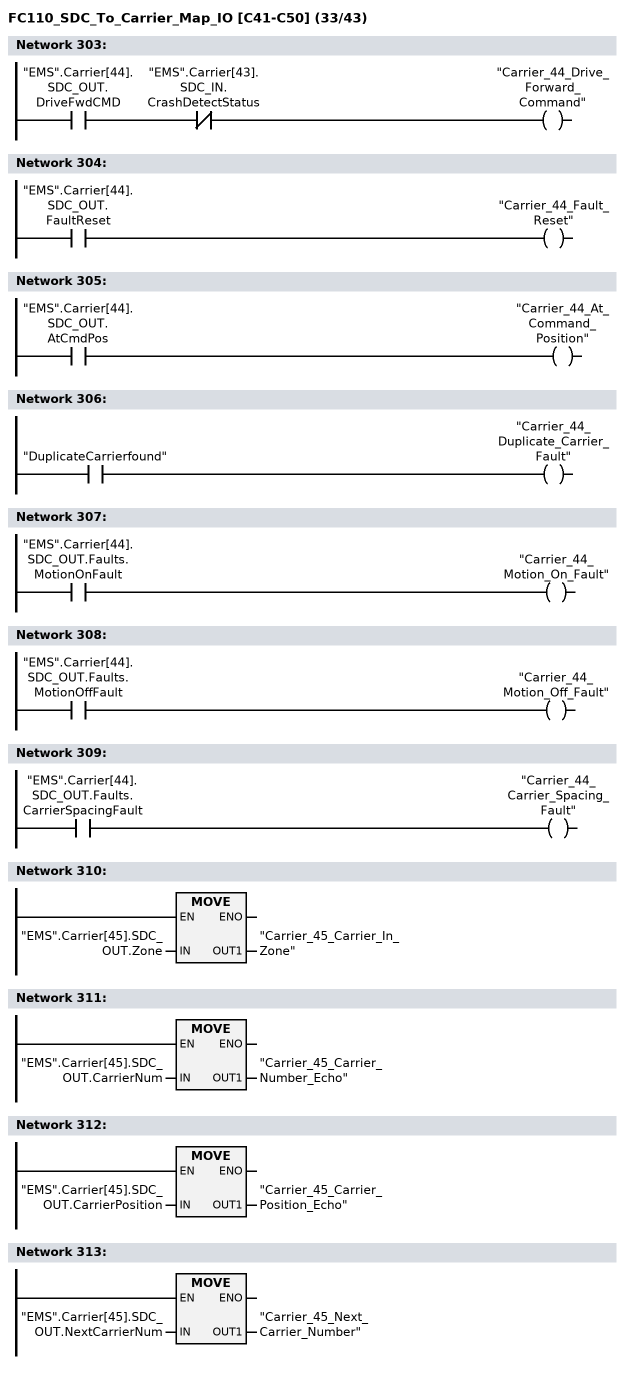
   RUNG wire#powerrail
      Contact( "EMS".Carrier[44].SDC_OUT.DriveFwdCMD )
      I_Contact( "EMS".Carrier[43].SDC_IN.CrashDetectStatus )
      Coil( "Carrier_44_Drive_Forward_Command" )
   END_RUNG
   // the same network as SCL:
   "Carrier_44_Drive_Forward_Command" := "EMS".Carrier[44].SDC_OUT.DriveFwdCMD AND NOT "EMS".Carrier[43].SDC_IN.CrashDetectStatus;
END_REGION

REGION Network 304
   RUNG wire#powerrail
      Contact( "EMS".Carrier[44].SDC_OUT.FaultReset )
      Coil( "Carrier_44_Fault_Reset" )
   END_RUNG
   // the same network as SCL:
   "Carrier_44_Fault_Reset" := "EMS".Carrier[44].SDC_OUT.FaultReset;
END_REGION

REGION Network 305
   RUNG wire#powerrail
      Contact( "EMS".Carrier[44].SDC_OUT.AtCmdPos )
      Coil( "Carrier_44_At_Command_Position" )
   END_RUNG
   // the same network as SCL:
   "Carrier_44_At_Command_Position" := "EMS".Carrier[44].SDC_OUT.AtCmdPos;
END_REGION

REGION Network 306
   RUNG wire#powerrail
      Contact( "DuplicateCarrierfound" )
      Coil( "Carrier_44_Duplicate_Carrier_Fault" )
   END_RUNG
   // the same network as SCL:
   "Carrier_44_Duplicate_Carrier_Fault" := "DuplicateCarrierfound";
END_REGION

REGION Network 307
   RUNG wire#powerrail
      Contact( "EMS".Carrier[44].SDC_OUT.Faults.MotionOnFault )
      Coil( "Carrier_44_Motion_On_Fault" )
   END_RUNG
   // the same network as SCL:
   "Carrier_44_Motion_On_Fault" := "EMS".Carrier[44].SDC_OUT.Faults.MotionOnFault;
END_REGION

REGION Network 308
   RUNG wire#powerrail
      Contact( "EMS".Carrier[44].SDC_OUT.Faults.MotionOffFault )
      Coil( "Carrier_44_Motion_Off_Fault" )
   END_RUNG
   // the same network as SCL:
   "Carrier_44_Motion_Off_Fault" := "EMS".Carrier[44].SDC_OUT.Faults.MotionOffFault;
END_REGION

REGION Network 309
   RUNG wire#powerrail
      Contact( "EMS".Carrier[44].SDC_OUT.Faults.CarrierSpacingFault )
      Coil( "Carrier_44_Carrier_Spacing_Fault" )
   END_RUNG
   // the same network as SCL:
   "Carrier_44_Carrier_Spacing_Fault" := "EMS".Carrier[44].SDC_OUT.Faults.CarrierSpacingFault;
END_REGION

REGION Network 310
   RUNG wire#powerrail
      Move(in := "EMS".Carrier[45].SDC_OUT.Zone, out1 => "Carrier_45_Carrier_In_Zone")
   END_RUNG
   // the same network as SCL:
   "Carrier_45_Carrier_In_Zone" := "EMS".Carrier[45].SDC_OUT.Zone;
END_REGION

REGION Network 311
   RUNG wire#powerrail
      Move(in := "EMS".Carrier[45].SDC_OUT.CarrierNum, out1 => "Carrier_45_Carrier_Number_Echo")
   END_RUNG
   // the same network as SCL:
   "Carrier_45_Carrier_Number_Echo" := "EMS".Carrier[45].SDC_OUT.CarrierNum;
END_REGION

REGION Network 312
   RUNG wire#powerrail
      Move(in := "EMS".Carrier[45].SDC_OUT.CarrierPosition, out1 => "Carrier_45_Carrier_Position_Echo")
   END_RUNG
   // the same network as SCL:
   "Carrier_45_Carrier_Position_Echo" := "EMS".Carrier[45].SDC_OUT.CarrierPosition;
END_REGION

REGION Network 313
   RUNG wire#powerrail
      Move(in := "EMS".Carrier[45].SDC_OUT.NextCarrierNum, out1 => "Carrier_45_Next_Carrier_Number")
   END_RUNG
   // the same network as SCL:
   "Carrier_45_Next_Carrier_Number" := "EMS".Carrier[45].SDC_OUT.NextCarrierNum;
END_REGION

REGION Network 314
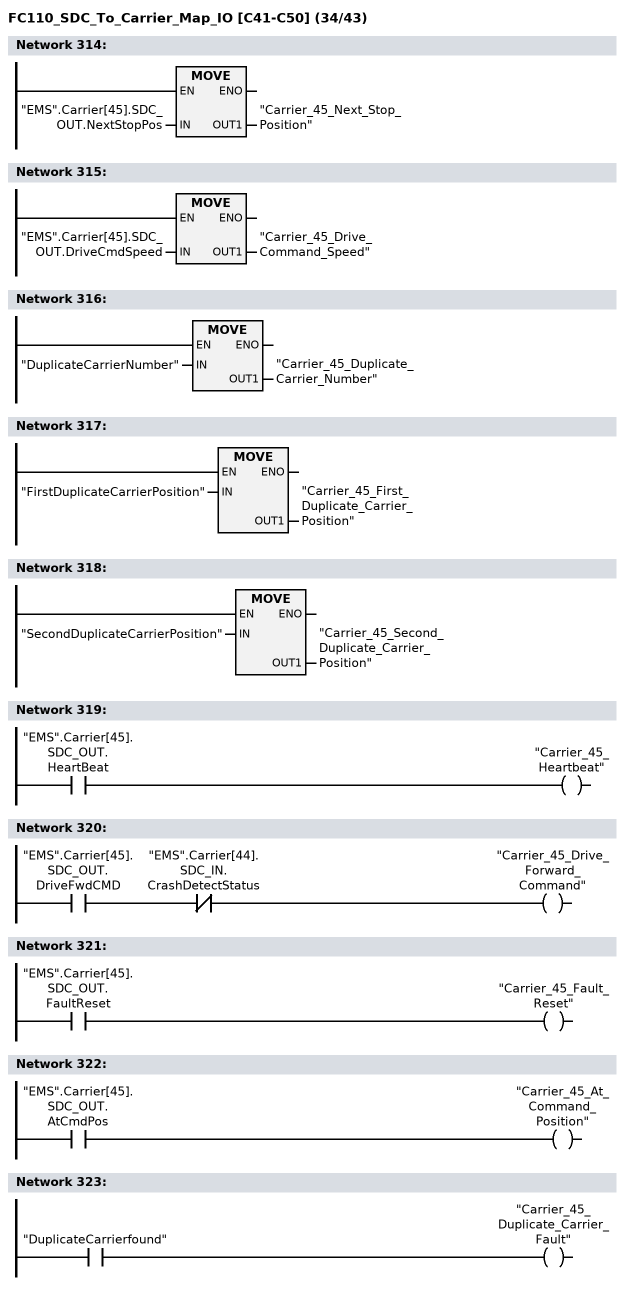
   RUNG wire#powerrail
      Move(in := "EMS".Carrier[45].SDC_OUT.NextStopPos, out1 => "Carrier_45_Next_Stop_Position")
   END_RUNG
   // the same network as SCL:
   "Carrier_45_Next_Stop_Position" := "EMS".Carrier[45].SDC_OUT.NextStopPos;
END_REGION

REGION Network 315
   RUNG wire#powerrail
      Move(in := "EMS".Carrier[45].SDC_OUT.DriveCmdSpeed, out1 => "Carrier_45_Drive_Command_Speed")
   END_RUNG
   // the same network as SCL:
   "Carrier_45_Drive_Command_Speed" := "EMS".Carrier[45].SDC_OUT.DriveCmdSpeed;
END_REGION

REGION Network 316
   RUNG wire#powerrail
      Move(in := "DuplicateCarrierNumber", out1 => "Carrier_45_Duplicate_Carrier_Number")
   END_RUNG
   // the same network as SCL:
   "Carrier_45_Duplicate_Carrier_Number" := "DuplicateCarrierNumber";
END_REGION

REGION Network 317
   RUNG wire#powerrail
      Move(in := "FirstDuplicateCarrierPosition", out1 => "Carrier_45_First_Duplicate_Carrier_Position")
   END_RUNG
   // the same network as SCL:
   "Carrier_45_First_Duplicate_Carrier_Position" := "FirstDuplicateCarrierPosition";
END_REGION

REGION Network 318
   RUNG wire#powerrail
      Move(in := "SecondDuplicateCarrierPosition", out1 => "Carrier_45_Second_Duplicate_Carrier_Position")
   END_RUNG
   // the same network as SCL:
   "Carrier_45_Second_Duplicate_Carrier_Position" := "SecondDuplicateCarrierPosition";
END_REGION

REGION Network 319
   RUNG wire#powerrail
      Contact( "EMS".Carrier[45].SDC_OUT.HeartBeat )
      Coil( "Carrier_45_Heartbeat" )
   END_RUNG
   // the same network as SCL:
   "Carrier_45_Heartbeat" := "EMS".Carrier[45].SDC_OUT.HeartBeat;
END_REGION

REGION Network 320
   RUNG wire#powerrail
      Contact( "EMS".Carrier[45].SDC_OUT.DriveFwdCMD )
      I_Contact( "EMS".Carrier[44].SDC_IN.CrashDetectStatus )
      Coil( "Carrier_45_Drive_Forward_Command" )
   END_RUNG
   // the same network as SCL:
   "Carrier_45_Drive_Forward_Command" := "EMS".Carrier[45].SDC_OUT.DriveFwdCMD AND NOT "EMS".Carrier[44].SDC_IN.CrashDetectStatus;
END_REGION

REGION Network 321
   RUNG wire#powerrail
      Contact( "EMS".Carrier[45].SDC_OUT.FaultReset )
      Coil( "Carrier_45_Fault_Reset" )
   END_RUNG
   // the same network as SCL:
   "Carrier_45_Fault_Reset" := "EMS".Carrier[45].SDC_OUT.FaultReset;
END_REGION

REGION Network 322
   RUNG wire#powerrail
      Contact( "EMS".Carrier[45].SDC_OUT.AtCmdPos )
      Coil( "Carrier_45_At_Command_Position" )
   END_RUNG
   // the same network as SCL:
   "Carrier_45_At_Command_Position" := "EMS".Carrier[45].SDC_OUT.AtCmdPos;
END_REGION

REGION Network 323
   RUNG wire#powerrail
      Contact( "DuplicateCarrierfound" )
      Coil( "Carrier_45_Duplicate_Carrier_Fault" )
   END_RUNG
   // the same network as SCL:
   "Carrier_45_Duplicate_Carrier_Fault" := "DuplicateCarrierfound";
END_REGION

REGION Network 324
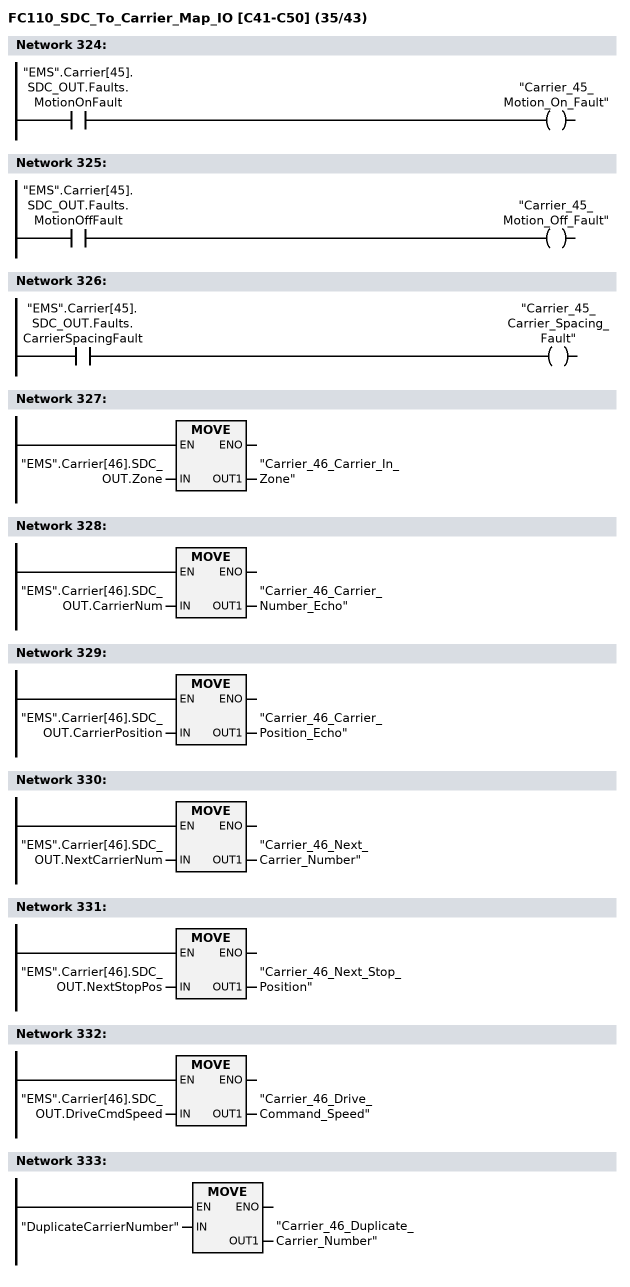
   RUNG wire#powerrail
      Contact( "EMS".Carrier[45].SDC_OUT.Faults.MotionOnFault )
      Coil( "Carrier_45_Motion_On_Fault" )
   END_RUNG
   // the same network as SCL:
   "Carrier_45_Motion_On_Fault" := "EMS".Carrier[45].SDC_OUT.Faults.MotionOnFault;
END_REGION

REGION Network 325
   RUNG wire#powerrail
      Contact( "EMS".Carrier[45].SDC_OUT.Faults.MotionOffFault )
      Coil( "Carrier_45_Motion_Off_Fault" )
   END_RUNG
   // the same network as SCL:
   "Carrier_45_Motion_Off_Fault" := "EMS".Carrier[45].SDC_OUT.Faults.MotionOffFault;
END_REGION

REGION Network 326
   RUNG wire#powerrail
      Contact( "EMS".Carrier[45].SDC_OUT.Faults.CarrierSpacingFault )
      Coil( "Carrier_45_Carrier_Spacing_Fault" )
   END_RUNG
   // the same network as SCL:
   "Carrier_45_Carrier_Spacing_Fault" := "EMS".Carrier[45].SDC_OUT.Faults.CarrierSpacingFault;
END_REGION

REGION Network 327
   RUNG wire#powerrail
      Move(in := "EMS".Carrier[46].SDC_OUT.Zone, out1 => "Carrier_46_Carrier_In_Zone")
   END_RUNG
   // the same network as SCL:
   "Carrier_46_Carrier_In_Zone" := "EMS".Carrier[46].SDC_OUT.Zone;
END_REGION

REGION Network 328
   RUNG wire#powerrail
      Move(in := "EMS".Carrier[46].SDC_OUT.CarrierNum, out1 => "Carrier_46_Carrier_Number_Echo")
   END_RUNG
   // the same network as SCL:
   "Carrier_46_Carrier_Number_Echo" := "EMS".Carrier[46].SDC_OUT.CarrierNum;
END_REGION

REGION Network 329
   RUNG wire#powerrail
      Move(in := "EMS".Carrier[46].SDC_OUT.CarrierPosition, out1 => "Carrier_46_Carrier_Position_Echo")
   END_RUNG
   // the same network as SCL:
   "Carrier_46_Carrier_Position_Echo" := "EMS".Carrier[46].SDC_OUT.CarrierPosition;
END_REGION

REGION Network 330
   RUNG wire#powerrail
      Move(in := "EMS".Carrier[46].SDC_OUT.NextCarrierNum, out1 => "Carrier_46_Next_Carrier_Number")
   END_RUNG
   // the same network as SCL:
   "Carrier_46_Next_Carrier_Number" := "EMS".Carrier[46].SDC_OUT.NextCarrierNum;
END_REGION

REGION Network 331
   RUNG wire#powerrail
      Move(in := "EMS".Carrier[46].SDC_OUT.NextStopPos, out1 => "Carrier_46_Next_Stop_Position")
   END_RUNG
   // the same network as SCL:
   "Carrier_46_Next_Stop_Position" := "EMS".Carrier[46].SDC_OUT.NextStopPos;
END_REGION

REGION Network 332
   RUNG wire#powerrail
      Move(in := "EMS".Carrier[46].SDC_OUT.DriveCmdSpeed, out1 => "Carrier_46_Drive_Command_Speed")
   END_RUNG
   // the same network as SCL:
   "Carrier_46_Drive_Command_Speed" := "EMS".Carrier[46].SDC_OUT.DriveCmdSpeed;
END_REGION

REGION Network 333
   RUNG wire#powerrail
      Move(in := "DuplicateCarrierNumber", out1 => "Carrier_46_Duplicate_Carrier_Number")
   END_RUNG
   // the same network as SCL:
   "Carrier_46_Duplicate_Carrier_Number" := "DuplicateCarrierNumber";
END_REGION

REGION Network 334
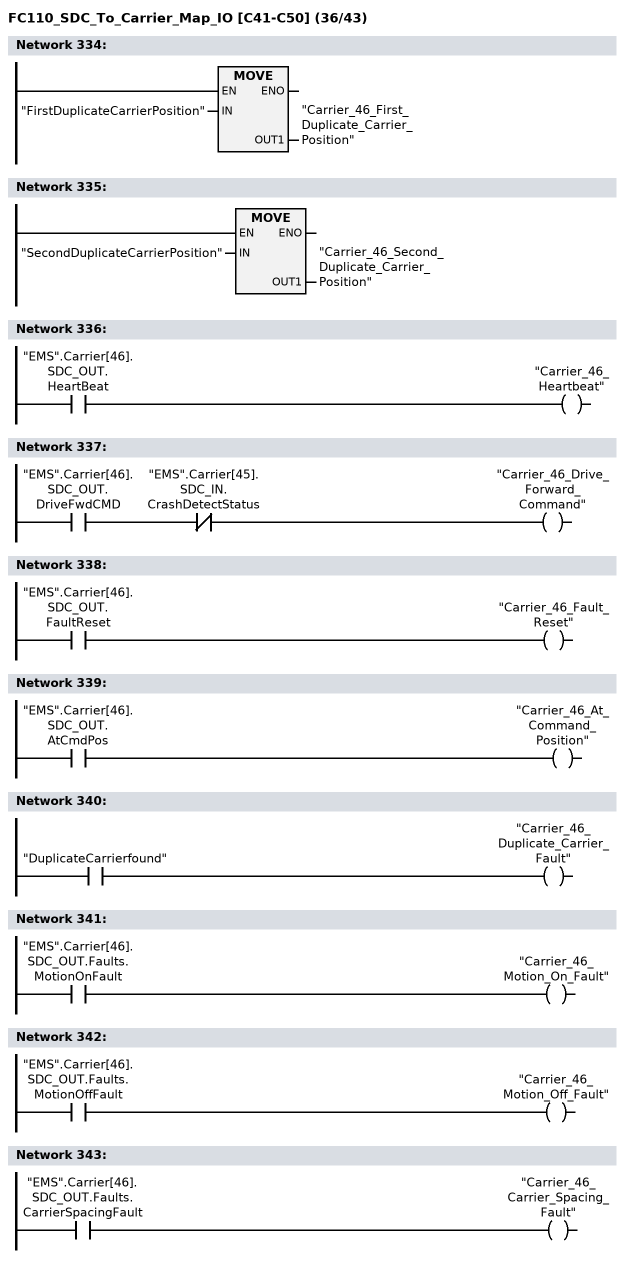
   RUNG wire#powerrail
      Move(in := "FirstDuplicateCarrierPosition", out1 => "Carrier_46_First_Duplicate_Carrier_Position")
   END_RUNG
   // the same network as SCL:
   "Carrier_46_First_Duplicate_Carrier_Position" := "FirstDuplicateCarrierPosition";
END_REGION

REGION Network 335
   RUNG wire#powerrail
      Move(in := "SecondDuplicateCarrierPosition", out1 => "Carrier_46_Second_Duplicate_Carrier_Position")
   END_RUNG
   // the same network as SCL:
   "Carrier_46_Second_Duplicate_Carrier_Position" := "SecondDuplicateCarrierPosition";
END_REGION

REGION Network 336
   RUNG wire#powerrail
      Contact( "EMS".Carrier[46].SDC_OUT.HeartBeat )
      Coil( "Carrier_46_Heartbeat" )
   END_RUNG
   // the same network as SCL:
   "Carrier_46_Heartbeat" := "EMS".Carrier[46].SDC_OUT.HeartBeat;
END_REGION

REGION Network 337
   RUNG wire#powerrail
      Contact( "EMS".Carrier[46].SDC_OUT.DriveFwdCMD )
      I_Contact( "EMS".Carrier[45].SDC_IN.CrashDetectStatus )
      Coil( "Carrier_46_Drive_Forward_Command" )
   END_RUNG
   // the same network as SCL:
   "Carrier_46_Drive_Forward_Command" := "EMS".Carrier[46].SDC_OUT.DriveFwdCMD AND NOT "EMS".Carrier[45].SDC_IN.CrashDetectStatus;
END_REGION

REGION Network 338
   RUNG wire#powerrail
      Contact( "EMS".Carrier[46].SDC_OUT.FaultReset )
      Coil( "Carrier_46_Fault_Reset" )
   END_RUNG
   // the same network as SCL:
   "Carrier_46_Fault_Reset" := "EMS".Carrier[46].SDC_OUT.FaultReset;
END_REGION

REGION Network 339
   RUNG wire#powerrail
      Contact( "EMS".Carrier[46].SDC_OUT.AtCmdPos )
      Coil( "Carrier_46_At_Command_Position" )
   END_RUNG
   // the same network as SCL:
   "Carrier_46_At_Command_Position" := "EMS".Carrier[46].SDC_OUT.AtCmdPos;
END_REGION

REGION Network 340
   RUNG wire#powerrail
      Contact( "DuplicateCarrierfound" )
      Coil( "Carrier_46_Duplicate_Carrier_Fault" )
   END_RUNG
   // the same network as SCL:
   "Carrier_46_Duplicate_Carrier_Fault" := "DuplicateCarrierfound";
END_REGION

REGION Network 341
   RUNG wire#powerrail
      Contact( "EMS".Carrier[46].SDC_OUT.Faults.MotionOnFault )
      Coil( "Carrier_46_Motion_On_Fault" )
   END_RUNG
   // the same network as SCL:
   "Carrier_46_Motion_On_Fault" := "EMS".Carrier[46].SDC_OUT.Faults.MotionOnFault;
END_REGION

REGION Network 342
   RUNG wire#powerrail
      Contact( "EMS".Carrier[46].SDC_OUT.Faults.MotionOffFault )
      Coil( "Carrier_46_Motion_Off_Fault" )
   END_RUNG
   // the same network as SCL:
   "Carrier_46_Motion_Off_Fault" := "EMS".Carrier[46].SDC_OUT.Faults.MotionOffFault;
END_REGION

REGION Network 343
   RUNG wire#powerrail
      Contact( "EMS".Carrier[46].SDC_OUT.Faults.CarrierSpacingFault )
      Coil( "Carrier_46_Carrier_Spacing_Fault" )
   END_RUNG
   // the same network as SCL:
   "Carrier_46_Carrier_Spacing_Fault" := "EMS".Carrier[46].SDC_OUT.Faults.CarrierSpacingFault;
END_REGION

REGION Network 344
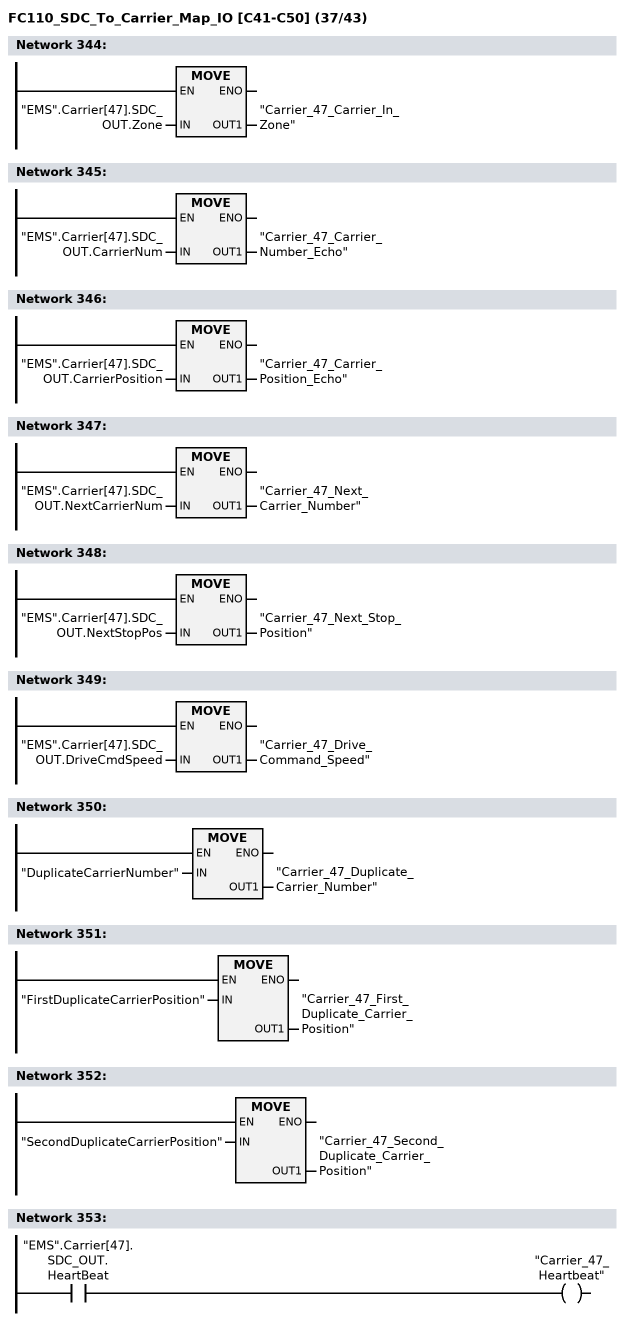
   RUNG wire#powerrail
      Move(in := "EMS".Carrier[47].SDC_OUT.Zone, out1 => "Carrier_47_Carrier_In_Zone")
   END_RUNG
   // the same network as SCL:
   "Carrier_47_Carrier_In_Zone" := "EMS".Carrier[47].SDC_OUT.Zone;
END_REGION

REGION Network 345
   RUNG wire#powerrail
      Move(in := "EMS".Carrier[47].SDC_OUT.CarrierNum, out1 => "Carrier_47_Carrier_Number_Echo")
   END_RUNG
   // the same network as SCL:
   "Carrier_47_Carrier_Number_Echo" := "EMS".Carrier[47].SDC_OUT.CarrierNum;
END_REGION

REGION Network 346
   RUNG wire#powerrail
      Move(in := "EMS".Carrier[47].SDC_OUT.CarrierPosition, out1 => "Carrier_47_Carrier_Position_Echo")
   END_RUNG
   // the same network as SCL:
   "Carrier_47_Carrier_Position_Echo" := "EMS".Carrier[47].SDC_OUT.CarrierPosition;
END_REGION

REGION Network 347
   RUNG wire#powerrail
      Move(in := "EMS".Carrier[47].SDC_OUT.NextCarrierNum, out1 => "Carrier_47_Next_Carrier_Number")
   END_RUNG
   // the same network as SCL:
   "Carrier_47_Next_Carrier_Number" := "EMS".Carrier[47].SDC_OUT.NextCarrierNum;
END_REGION

REGION Network 348
   RUNG wire#powerrail
      Move(in := "EMS".Carrier[47].SDC_OUT.NextStopPos, out1 => "Carrier_47_Next_Stop_Position")
   END_RUNG
   // the same network as SCL:
   "Carrier_47_Next_Stop_Position" := "EMS".Carrier[47].SDC_OUT.NextStopPos;
END_REGION

REGION Network 349
   RUNG wire#powerrail
      Move(in := "EMS".Carrier[47].SDC_OUT.DriveCmdSpeed, out1 => "Carrier_47_Drive_Command_Speed")
   END_RUNG
   // the same network as SCL:
   "Carrier_47_Drive_Command_Speed" := "EMS".Carrier[47].SDC_OUT.DriveCmdSpeed;
END_REGION

REGION Network 350
   RUNG wire#powerrail
      Move(in := "DuplicateCarrierNumber", out1 => "Carrier_47_Duplicate_Carrier_Number")
   END_RUNG
   // the same network as SCL:
   "Carrier_47_Duplicate_Carrier_Number" := "DuplicateCarrierNumber";
END_REGION

REGION Network 351
   RUNG wire#powerrail
      Move(in := "FirstDuplicateCarrierPosition", out1 => "Carrier_47_First_Duplicate_Carrier_Position")
   END_RUNG
   // the same network as SCL:
   "Carrier_47_First_Duplicate_Carrier_Position" := "FirstDuplicateCarrierPosition";
END_REGION

REGION Network 352
   RUNG wire#powerrail
      Move(in := "SecondDuplicateCarrierPosition", out1 => "Carrier_47_Second_Duplicate_Carrier_Position")
   END_RUNG
   // the same network as SCL:
   "Carrier_47_Second_Duplicate_Carrier_Position" := "SecondDuplicateCarrierPosition";
END_REGION

REGION Network 353
   RUNG wire#powerrail
      Contact( "EMS".Carrier[47].SDC_OUT.HeartBeat )
      Coil( "Carrier_47_Heartbeat" )
   END_RUNG
   // the same network as SCL:
   "Carrier_47_Heartbeat" := "EMS".Carrier[47].SDC_OUT.HeartBeat;
END_REGION

REGION Network 354
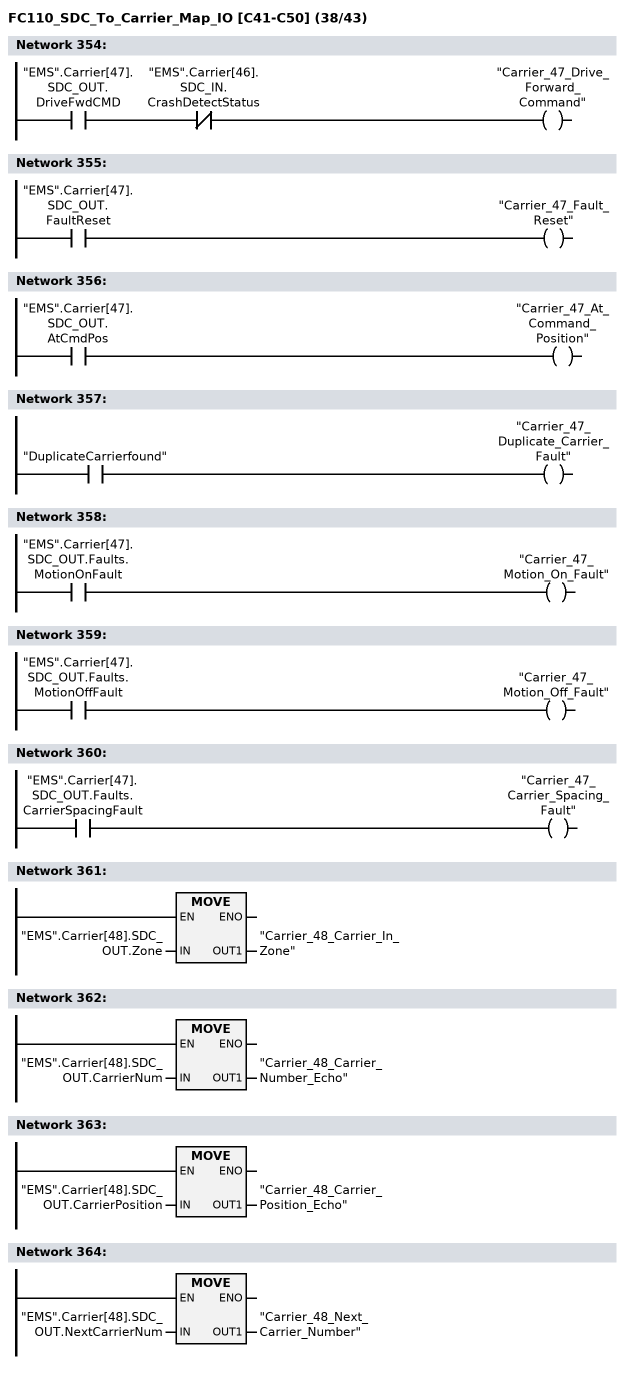
   RUNG wire#powerrail
      Contact( "EMS".Carrier[47].SDC_OUT.DriveFwdCMD )
      I_Contact( "EMS".Carrier[46].SDC_IN.CrashDetectStatus )
      Coil( "Carrier_47_Drive_Forward_Command" )
   END_RUNG
   // the same network as SCL:
   "Carrier_47_Drive_Forward_Command" := "EMS".Carrier[47].SDC_OUT.DriveFwdCMD AND NOT "EMS".Carrier[46].SDC_IN.CrashDetectStatus;
END_REGION

REGION Network 355
   RUNG wire#powerrail
      Contact( "EMS".Carrier[47].SDC_OUT.FaultReset )
      Coil( "Carrier_47_Fault_Reset" )
   END_RUNG
   // the same network as SCL:
   "Carrier_47_Fault_Reset" := "EMS".Carrier[47].SDC_OUT.FaultReset;
END_REGION

REGION Network 356
   RUNG wire#powerrail
      Contact( "EMS".Carrier[47].SDC_OUT.AtCmdPos )
      Coil( "Carrier_47_At_Command_Position" )
   END_RUNG
   // the same network as SCL:
   "Carrier_47_At_Command_Position" := "EMS".Carrier[47].SDC_OUT.AtCmdPos;
END_REGION

REGION Network 357
   RUNG wire#powerrail
      Contact( "DuplicateCarrierfound" )
      Coil( "Carrier_47_Duplicate_Carrier_Fault" )
   END_RUNG
   // the same network as SCL:
   "Carrier_47_Duplicate_Carrier_Fault" := "DuplicateCarrierfound";
END_REGION

REGION Network 358
   RUNG wire#powerrail
      Contact( "EMS".Carrier[47].SDC_OUT.Faults.MotionOnFault )
      Coil( "Carrier_47_Motion_On_Fault" )
   END_RUNG
   // the same network as SCL:
   "Carrier_47_Motion_On_Fault" := "EMS".Carrier[47].SDC_OUT.Faults.MotionOnFault;
END_REGION

REGION Network 359
   RUNG wire#powerrail
      Contact( "EMS".Carrier[47].SDC_OUT.Faults.MotionOffFault )
      Coil( "Carrier_47_Motion_Off_Fault" )
   END_RUNG
   // the same network as SCL:
   "Carrier_47_Motion_Off_Fault" := "EMS".Carrier[47].SDC_OUT.Faults.MotionOffFault;
END_REGION

REGION Network 360
   RUNG wire#powerrail
      Contact( "EMS".Carrier[47].SDC_OUT.Faults.CarrierSpacingFault )
      Coil( "Carrier_47_Carrier_Spacing_Fault" )
   END_RUNG
   // the same network as SCL:
   "Carrier_47_Carrier_Spacing_Fault" := "EMS".Carrier[47].SDC_OUT.Faults.CarrierSpacingFault;
END_REGION

REGION Network 361
   RUNG wire#powerrail
      Move(in := "EMS".Carrier[48].SDC_OUT.Zone, out1 => "Carrier_48_Carrier_In_Zone")
   END_RUNG
   // the same network as SCL:
   "Carrier_48_Carrier_In_Zone" := "EMS".Carrier[48].SDC_OUT.Zone;
END_REGION

REGION Network 362
   RUNG wire#powerrail
      Move(in := "EMS".Carrier[48].SDC_OUT.CarrierNum, out1 => "Carrier_48_Carrier_Number_Echo")
   END_RUNG
   // the same network as SCL:
   "Carrier_48_Carrier_Number_Echo" := "EMS".Carrier[48].SDC_OUT.CarrierNum;
END_REGION

REGION Network 363
   RUNG wire#powerrail
      Move(in := "EMS".Carrier[48].SDC_OUT.CarrierPosition, out1 => "Carrier_48_Carrier_Position_Echo")
   END_RUNG
   // the same network as SCL:
   "Carrier_48_Carrier_Position_Echo" := "EMS".Carrier[48].SDC_OUT.CarrierPosition;
END_REGION

REGION Network 364
   RUNG wire#powerrail
      Move(in := "EMS".Carrier[48].SDC_OUT.NextCarrierNum, out1 => "Carrier_48_Next_Carrier_Number")
   END_RUNG
   // the same network as SCL:
   "Carrier_48_Next_Carrier_Number" := "EMS".Carrier[48].SDC_OUT.NextCarrierNum;
END_REGION

REGION Network 365
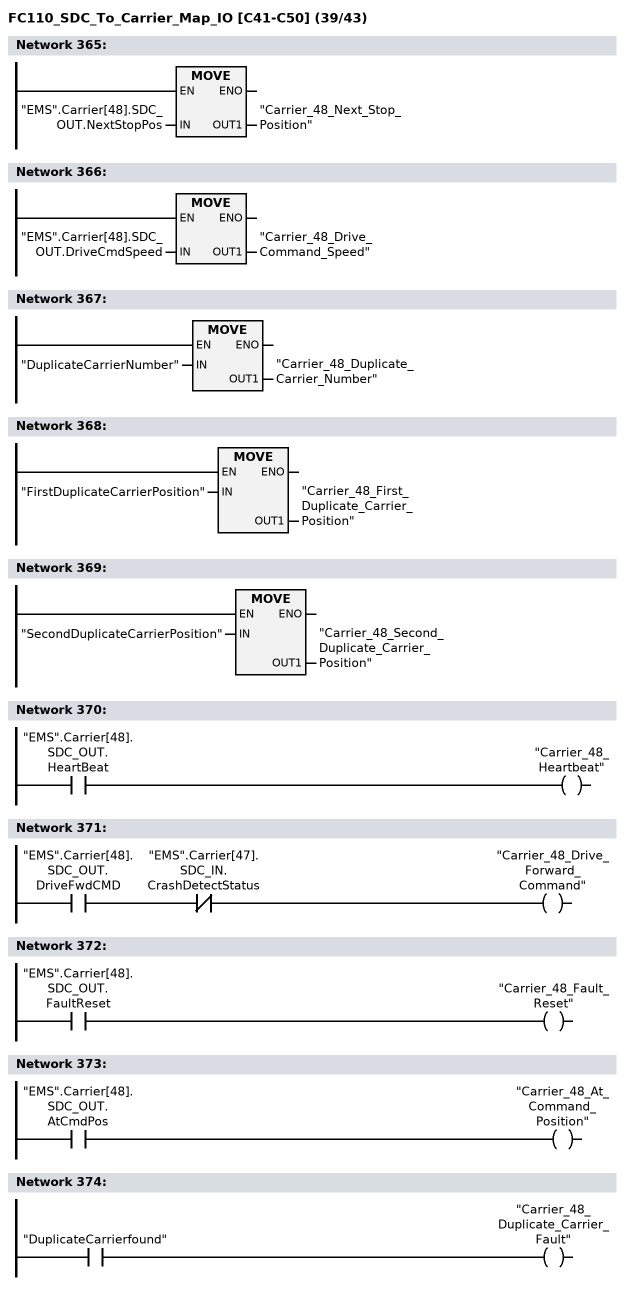
   RUNG wire#powerrail
      Move(in := "EMS".Carrier[48].SDC_OUT.NextStopPos, out1 => "Carrier_48_Next_Stop_Position")
   END_RUNG
   // the same network as SCL:
   "Carrier_48_Next_Stop_Position" := "EMS".Carrier[48].SDC_OUT.NextStopPos;
END_REGION

REGION Network 366
   RUNG wire#powerrail
      Move(in := "EMS".Carrier[48].SDC_OUT.DriveCmdSpeed, out1 => "Carrier_48_Drive_Command_Speed")
   END_RUNG
   // the same network as SCL:
   "Carrier_48_Drive_Command_Speed" := "EMS".Carrier[48].SDC_OUT.DriveCmdSpeed;
END_REGION

REGION Network 367
   RUNG wire#powerrail
      Move(in := "DuplicateCarrierNumber", out1 => "Carrier_48_Duplicate_Carrier_Number")
   END_RUNG
   // the same network as SCL:
   "Carrier_48_Duplicate_Carrier_Number" := "DuplicateCarrierNumber";
END_REGION

REGION Network 368
   RUNG wire#powerrail
      Move(in := "FirstDuplicateCarrierPosition", out1 => "Carrier_48_First_Duplicate_Carrier_Position")
   END_RUNG
   // the same network as SCL:
   "Carrier_48_First_Duplicate_Carrier_Position" := "FirstDuplicateCarrierPosition";
END_REGION

REGION Network 369
   RUNG wire#powerrail
      Move(in := "SecondDuplicateCarrierPosition", out1 => "Carrier_48_Second_Duplicate_Carrier_Position")
   END_RUNG
   // the same network as SCL:
   "Carrier_48_Second_Duplicate_Carrier_Position" := "SecondDuplicateCarrierPosition";
END_REGION

REGION Network 370
   RUNG wire#powerrail
      Contact( "EMS".Carrier[48].SDC_OUT.HeartBeat )
      Coil( "Carrier_48_Heartbeat" )
   END_RUNG
   // the same network as SCL:
   "Carrier_48_Heartbeat" := "EMS".Carrier[48].SDC_OUT.HeartBeat;
END_REGION

REGION Network 371
   RUNG wire#powerrail
      Contact( "EMS".Carrier[48].SDC_OUT.DriveFwdCMD )
      I_Contact( "EMS".Carrier[47].SDC_IN.CrashDetectStatus )
      Coil( "Carrier_48_Drive_Forward_Command" )
   END_RUNG
   // the same network as SCL:
   "Carrier_48_Drive_Forward_Command" := "EMS".Carrier[48].SDC_OUT.DriveFwdCMD AND NOT "EMS".Carrier[47].SDC_IN.CrashDetectStatus;
END_REGION

REGION Network 372
   RUNG wire#powerrail
      Contact( "EMS".Carrier[48].SDC_OUT.FaultReset )
      Coil( "Carrier_48_Fault_Reset" )
   END_RUNG
   // the same network as SCL:
   "Carrier_48_Fault_Reset" := "EMS".Carrier[48].SDC_OUT.FaultReset;
END_REGION

REGION Network 373
   RUNG wire#powerrail
      Contact( "EMS".Carrier[48].SDC_OUT.AtCmdPos )
      Coil( "Carrier_48_At_Command_Position" )
   END_RUNG
   // the same network as SCL:
   "Carrier_48_At_Command_Position" := "EMS".Carrier[48].SDC_OUT.AtCmdPos;
END_REGION

REGION Network 374
   RUNG wire#powerrail
      Contact( "DuplicateCarrierfound" )
      Coil( "Carrier_48_Duplicate_Carrier_Fault" )
   END_RUNG
   // the same network as SCL:
   "Carrier_48_Duplicate_Carrier_Fault" := "DuplicateCarrierfound";
END_REGION

REGION Network 375
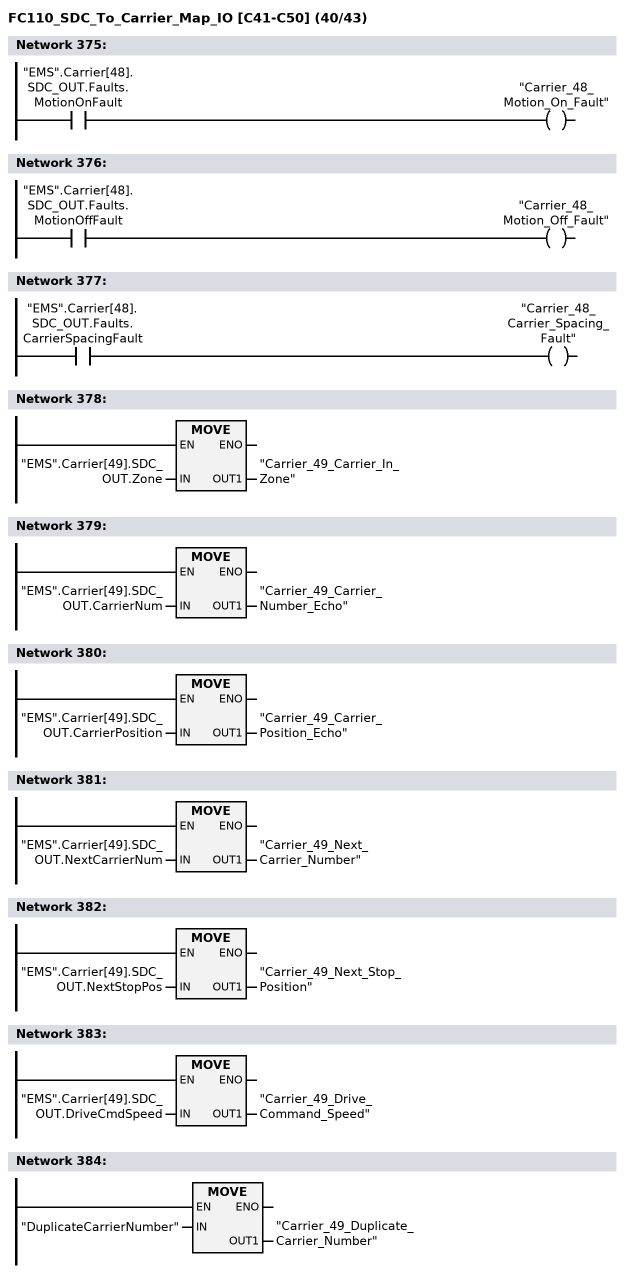
   RUNG wire#powerrail
      Contact( "EMS".Carrier[48].SDC_OUT.Faults.MotionOnFault )
      Coil( "Carrier_48_Motion_On_Fault" )
   END_RUNG
   // the same network as SCL:
   "Carrier_48_Motion_On_Fault" := "EMS".Carrier[48].SDC_OUT.Faults.MotionOnFault;
END_REGION

REGION Network 376
   RUNG wire#powerrail
      Contact( "EMS".Carrier[48].SDC_OUT.Faults.MotionOffFault )
      Coil( "Carrier_48_Motion_Off_Fault" )
   END_RUNG
   // the same network as SCL:
   "Carrier_48_Motion_Off_Fault" := "EMS".Carrier[48].SDC_OUT.Faults.MotionOffFault;
END_REGION

REGION Network 377
   RUNG wire#powerrail
      Contact( "EMS".Carrier[48].SDC_OUT.Faults.CarrierSpacingFault )
      Coil( "Carrier_48_Carrier_Spacing_Fault" )
   END_RUNG
   // the same network as SCL:
   "Carrier_48_Carrier_Spacing_Fault" := "EMS".Carrier[48].SDC_OUT.Faults.CarrierSpacingFault;
END_REGION

REGION Network 378
   RUNG wire#powerrail
      Move(in := "EMS".Carrier[49].SDC_OUT.Zone, out1 => "Carrier_49_Carrier_In_Zone")
   END_RUNG
   // the same network as SCL:
   "Carrier_49_Carrier_In_Zone" := "EMS".Carrier[49].SDC_OUT.Zone;
END_REGION

REGION Network 379
   RUNG wire#powerrail
      Move(in := "EMS".Carrier[49].SDC_OUT.CarrierNum, out1 => "Carrier_49_Carrier_Number_Echo")
   END_RUNG
   // the same network as SCL:
   "Carrier_49_Carrier_Number_Echo" := "EMS".Carrier[49].SDC_OUT.CarrierNum;
END_REGION

REGION Network 380
   RUNG wire#powerrail
      Move(in := "EMS".Carrier[49].SDC_OUT.CarrierPosition, out1 => "Carrier_49_Carrier_Position_Echo")
   END_RUNG
   // the same network as SCL:
   "Carrier_49_Carrier_Position_Echo" := "EMS".Carrier[49].SDC_OUT.CarrierPosition;
END_REGION

REGION Network 381
   RUNG wire#powerrail
      Move(in := "EMS".Carrier[49].SDC_OUT.NextCarrierNum, out1 => "Carrier_49_Next_Carrier_Number")
   END_RUNG
   // the same network as SCL:
   "Carrier_49_Next_Carrier_Number" := "EMS".Carrier[49].SDC_OUT.NextCarrierNum;
END_REGION

REGION Network 382
   RUNG wire#powerrail
      Move(in := "EMS".Carrier[49].SDC_OUT.NextStopPos, out1 => "Carrier_49_Next_Stop_Position")
   END_RUNG
   // the same network as SCL:
   "Carrier_49_Next_Stop_Position" := "EMS".Carrier[49].SDC_OUT.NextStopPos;
END_REGION

REGION Network 383
   RUNG wire#powerrail
      Move(in := "EMS".Carrier[49].SDC_OUT.DriveCmdSpeed, out1 => "Carrier_49_Drive_Command_Speed")
   END_RUNG
   // the same network as SCL:
   "Carrier_49_Drive_Command_Speed" := "EMS".Carrier[49].SDC_OUT.DriveCmdSpeed;
END_REGION

REGION Network 384
   RUNG wire#powerrail
      Move(in := "DuplicateCarrierNumber", out1 => "Carrier_49_Duplicate_Carrier_Number")
   END_RUNG
   // the same network as SCL:
   "Carrier_49_Duplicate_Carrier_Number" := "DuplicateCarrierNumber";
END_REGION

REGION Network 385
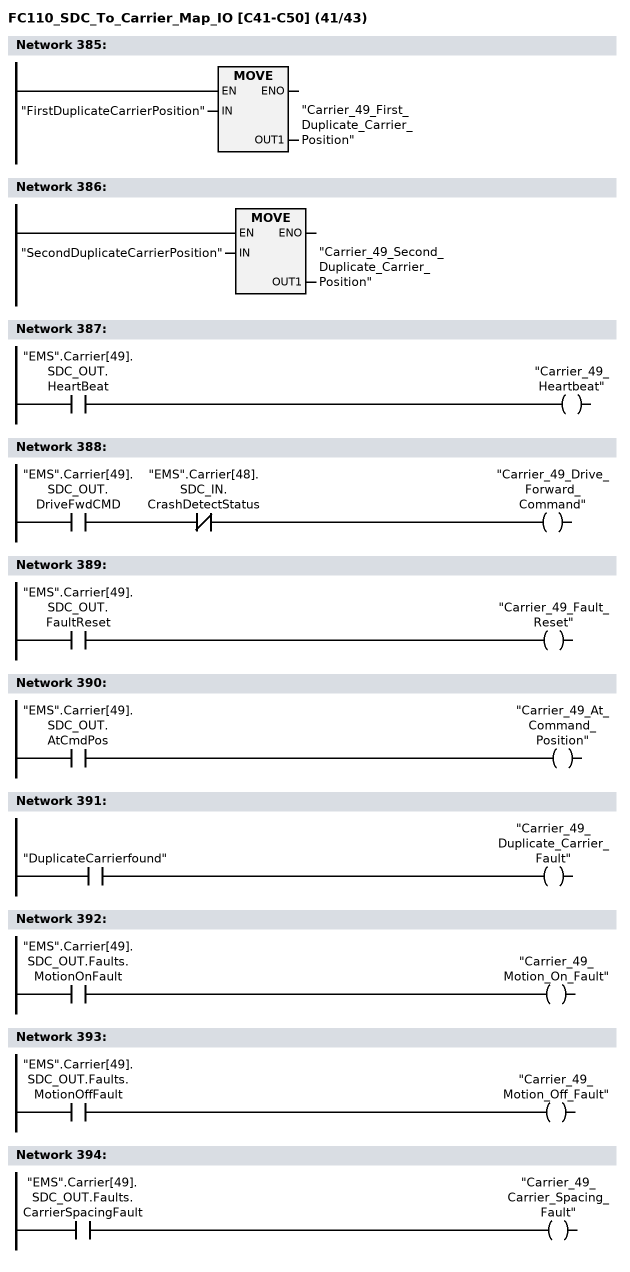
   RUNG wire#powerrail
      Move(in := "FirstDuplicateCarrierPosition", out1 => "Carrier_49_First_Duplicate_Carrier_Position")
   END_RUNG
   // the same network as SCL:
   "Carrier_49_First_Duplicate_Carrier_Position" := "FirstDuplicateCarrierPosition";
END_REGION

REGION Network 386
   RUNG wire#powerrail
      Move(in := "SecondDuplicateCarrierPosition", out1 => "Carrier_49_Second_Duplicate_Carrier_Position")
   END_RUNG
   // the same network as SCL:
   "Carrier_49_Second_Duplicate_Carrier_Position" := "SecondDuplicateCarrierPosition";
END_REGION

REGION Network 387
   RUNG wire#powerrail
      Contact( "EMS".Carrier[49].SDC_OUT.HeartBeat )
      Coil( "Carrier_49_Heartbeat" )
   END_RUNG
   // the same network as SCL:
   "Carrier_49_Heartbeat" := "EMS".Carrier[49].SDC_OUT.HeartBeat;
END_REGION

REGION Network 388
   RUNG wire#powerrail
      Contact( "EMS".Carrier[49].SDC_OUT.DriveFwdCMD )
      I_Contact( "EMS".Carrier[48].SDC_IN.CrashDetectStatus )
      Coil( "Carrier_49_Drive_Forward_Command" )
   END_RUNG
   // the same network as SCL:
   "Carrier_49_Drive_Forward_Command" := "EMS".Carrier[49].SDC_OUT.DriveFwdCMD AND NOT "EMS".Carrier[48].SDC_IN.CrashDetectStatus;
END_REGION

REGION Network 389
   RUNG wire#powerrail
      Contact( "EMS".Carrier[49].SDC_OUT.FaultReset )
      Coil( "Carrier_49_Fault_Reset" )
   END_RUNG
   // the same network as SCL:
   "Carrier_49_Fault_Reset" := "EMS".Carrier[49].SDC_OUT.FaultReset;
END_REGION

REGION Network 390
   RUNG wire#powerrail
      Contact( "EMS".Carrier[49].SDC_OUT.AtCmdPos )
      Coil( "Carrier_49_At_Command_Position" )
   END_RUNG
   // the same network as SCL:
   "Carrier_49_At_Command_Position" := "EMS".Carrier[49].SDC_OUT.AtCmdPos;
END_REGION

REGION Network 391
   RUNG wire#powerrail
      Contact( "DuplicateCarrierfound" )
      Coil( "Carrier_49_Duplicate_Carrier_Fault" )
   END_RUNG
   // the same network as SCL:
   "Carrier_49_Duplicate_Carrier_Fault" := "DuplicateCarrierfound";
END_REGION

REGION Network 392
   RUNG wire#powerrail
      Contact( "EMS".Carrier[49].SDC_OUT.Faults.MotionOnFault )
      Coil( "Carrier_49_Motion_On_Fault" )
   END_RUNG
   // the same network as SCL:
   "Carrier_49_Motion_On_Fault" := "EMS".Carrier[49].SDC_OUT.Faults.MotionOnFault;
END_REGION

REGION Network 393
   RUNG wire#powerrail
      Contact( "EMS".Carrier[49].SDC_OUT.Faults.MotionOffFault )
      Coil( "Carrier_49_Motion_Off_Fault" )
   END_RUNG
   // the same network as SCL:
   "Carrier_49_Motion_Off_Fault" := "EMS".Carrier[49].SDC_OUT.Faults.MotionOffFault;
END_REGION

REGION Network 394
   RUNG wire#powerrail
      Contact( "EMS".Carrier[49].SDC_OUT.Faults.CarrierSpacingFault )
      Coil( "Carrier_49_Carrier_Spacing_Fault" )
   END_RUNG
   // the same network as SCL:
   "Carrier_49_Carrier_Spacing_Fault" := "EMS".Carrier[49].SDC_OUT.Faults.CarrierSpacingFault;
END_REGION

REGION Network 395
